(* Logix 5000 project; controller MV vendor 1 type 14 code 217 rev 31.11; software revision 31.00; part 49 of 53 *)
(* tags used below, declared in another part *)
   CheckTimeMask : INT;
   CWD : CHECKWORD_FLAGS;
   Delphi_Does_Eng_Func : BOOL;
   MV_MV10R : PlantItem;   // MV10R
   MV_MV11R : PlantItem;   // MV11R
   MV_MV12R : PlantItem;   // MV12R
   MV_MV13R : PlantItem;   // MV13R
   MV_MV14R : PlantItem;   // MV14R
   MV_MV15R : PlantItem;   // MV15R
   MV_MV16R : PlantItem;   // MV16R
   MV_MV17R : PlantItem;   // MV17R
   MV_MV18R : PlantItem;   // MV18R
   MV_MV19R : PlantItem;   // MV19R
   MV_MV1R : PlantItem;   // MV1R
   MV_MV20R : PlantItem;   // MV20R
   MV_MV21R : PlantItem;   // MV21R
   MV_MV22R : PlantItem;   // MV22R
   MV_MV23R : PlantItem;   // MV23R
   MV_MV2R : PlantItem;   // MV2R
   MV_MV30R : PlantItem;   // MV30R
   MV_MV31R : PlantItem;   // MV31R
   MV_MV32R : PlantItem;   // MV32R
   MV_MV33R : PlantItem;   // MV33R
   MV_MV34R : PlantItem;   // MV34R
   MV_MV35R : PlantItem;   // MV35R
   MV_MV3R : PlantItem;   // MV3R
   MV_MV4R : PlantItem;   // MV4R
   MV_MV5R : PlantItem;   // MV5R
   MV_MV6R : PlantItem;   // MV6R
   MV_MV8R : PlantItem;   // MV8R
   MV_MV9R : PlantItem;   // MV9R
   MV_N255 : DINT[255];   // Old Format Checkwords To Keep Delphi Indicating Status Correctly.
   TempChecktime : DINT;
(* MV_Common, continued *)

   48: [XIC(Delphi_Does_Eng_Func) [[XIC(MV_N255[39].8) [OTL(MV_MV8R.CW.[CWD.MANUAL]) ,XIC(MV_N255[39].9) OTL(MV_MV8R.CW.[CWD.MANDRV]) ,XIO(MV_N255[39].9) OTU(MV_MV8R.CW.[CWD.MANDRV]) ] ,XIO(MV_N255[39].8) [OTU(MV_MV8R.CW.[CWD.MANUAL]) ,[XIC(MV_MV8R.CW.[CWD.OUTPUT]) OTL(MV_N255[39].9) ,XIO(MV_MV8R.CW.[CWD.OUTPUT]) OTU(MV_N255[39].9) ] ] ] ,[XIC(MV_N255[39].13) OTL(MV_MV8R.CW.[CWD.CHECKOFF]) ,XIO(MV_N255[39].13) OTU(MV_MV8R.CW.[CWD.CHECKOFF]) ] ] ,XIO(Delphi_Does_Eng_Func) [[XIC(MV_MV8R.CW.[CWD.MANUAL]) OTL(MV_N255[39].8) ,XIO(MV_MV8R.CW.[CWD.MANUAL]) OTU(MV_N255[39].8) ] ,[XIC(MV_MV8R.CW.[CWD.CHECKOFF]) OTL(MV_N255[39].13) ,XIO(MV_MV8R.CW.[CWD.CHECKOFF]) OTU(MV_N255[39].13) ] ,[XIC(MV_MV8R.CW.[CWD.OUTPUT]) OTL(MV_N255[39].9) ,XIO(MV_MV8R.CW.[CWD.OUTPUT]) OTU(MV_N255[39].9) ] ] ,XIC(MV_MV8R.CW.[CWD.RUNFB]) OTE(MV_N255[39].10) ,XIO(MV_MV8R.CW.[CWD.RUNFB]) OTE(MV_N255[39].11) ,XIC(MV_MV8R.CW.[CWD.FAULT]) OTE(MV_N255[39].15) ];
   49: [XIC(Delphi_Does_Eng_Func) [[XIC(MV_N255[40].8) [OTL(MV_MV9R.CW.[CWD.MANUAL]) ,XIC(MV_N255[40].9) OTL(MV_MV9R.CW.[CWD.MANDRV]) ,XIO(MV_N255[40].9) OTU(MV_MV9R.CW.[CWD.MANDRV]) ] ,XIO(MV_N255[40].8) [OTU(MV_MV9R.CW.[CWD.MANUAL]) ,[XIC(MV_MV9R.CW.[CWD.OUTPUT]) OTL(MV_N255[40].9) ,XIO(MV_MV9R.CW.[CWD.OUTPUT]) OTU(MV_N255[40].9) ] ] ] ,[XIC(MV_N255[40].13) OTL(MV_MV9R.CW.[CWD.CHECKOFF]) ,XIO(MV_N255[40].13) OTU(MV_MV9R.CW.[CWD.CHECKOFF]) ] ] ,XIO(Delphi_Does_Eng_Func) [[XIC(MV_MV9R.CW.[CWD.MANUAL]) OTL(MV_N255[40].8) ,XIO(MV_MV9R.CW.[CWD.MANUAL]) OTU(MV_N255[40].8) ] ,[XIC(MV_MV9R.CW.[CWD.CHECKOFF]) OTL(MV_N255[40].13) ,XIO(MV_MV9R.CW.[CWD.CHECKOFF]) OTU(MV_N255[40].13) ] ,[XIC(MV_MV9R.CW.[CWD.OUTPUT]) OTL(MV_N255[40].9) ,XIO(MV_MV9R.CW.[CWD.OUTPUT]) OTU(MV_N255[40].9) ] ] ,XIC(MV_MV9R.CW.[CWD.RUNFB]) OTE(MV_N255[40].10) ,XIO(MV_MV9R.CW.[CWD.RUNFB]) OTE(MV_N255[40].11) ,XIC(MV_MV9R.CW.[CWD.FAULT]) OTE(MV_N255[40].15) ];
   50: [XIC(Delphi_Does_Eng_Func) [[XIC(MV_N255[41].8) [OTL(MV_MV10R.CW.[CWD.MANUAL]) ,XIC(MV_N255[41].9) OTL(MV_MV10R.CW.[CWD.MANDRV]) ,XIO(MV_N255[41].9) OTU(MV_MV10R.CW.[CWD.MANDRV]) ] ,XIO(MV_N255[41].8) [OTU(MV_MV10R.CW.[CWD.MANUAL]) ,[XIC(MV_MV10R.CW.[CWD.OUTPUT]) OTL(MV_N255[41].9) ,XIO(MV_MV10R.CW.[CWD.OUTPUT]) OTU(MV_N255[41].9) ] ] ] ,[XIC(MV_N255[41].13) OTL(MV_MV10R.CW.[CWD.CHECKOFF]) ,XIO(MV_N255[41].13) OTU(MV_MV10R.CW.[CWD.CHECKOFF]) ] ] ,XIO(Delphi_Does_Eng_Func) [[XIC(MV_MV10R.CW.[CWD.MANUAL]) OTL(MV_N255[41].8) ,XIO(MV_MV10R.CW.[CWD.MANUAL]) OTU(MV_N255[41].8) ] ,[XIC(MV_MV10R.CW.[CWD.CHECKOFF]) OTL(MV_N255[41].13) ,XIO(MV_MV10R.CW.[CWD.CHECKOFF]) OTU(MV_N255[41].13) ] ,[XIC(MV_MV10R.CW.[CWD.OUTPUT]) OTL(MV_N255[41].9) ,XIO(MV_MV10R.CW.[CWD.OUTPUT]) OTU(MV_N255[41].9) ] ] ,XIC(MV_MV10R.CW.[CWD.RUNFB]) OTE(MV_N255[41].10) ,XIO(MV_MV10R.CW.[CWD.RUNFB]) OTE(MV_N255[41].11) ,XIC(MV_MV10R.CW.[CWD.FAULT]) OTE(MV_N255[41].15) ];
   51: [XIC(Delphi_Does_Eng_Func) [[XIC(MV_N255[42].8) [OTL(MV_MV11R.CW.[CWD.MANUAL]) ,XIC(MV_N255[42].9) OTL(MV_MV11R.CW.[CWD.MANDRV]) ,XIO(MV_N255[42].9) OTU(MV_MV11R.CW.[CWD.MANDRV]) ] ,XIO(MV_N255[42].8) [OTU(MV_MV11R.CW.[CWD.MANUAL]) ,[XIC(MV_MV11R.CW.[CWD.OUTPUT]) OTL(MV_N255[42].9) ,XIO(MV_MV11R.CW.[CWD.OUTPUT]) OTU(MV_N255[42].9) ] ] ] ,[XIC(MV_N255[42].13) OTL(MV_MV11R.CW.[CWD.CHECKOFF]) ,XIO(MV_N255[42].13) OTU(MV_MV11R.CW.[CWD.CHECKOFF]) ] ] ,XIO(Delphi_Does_Eng_Func) [[XIC(MV_MV11R.CW.[CWD.MANUAL]) OTL(MV_N255[42].8) ,XIO(MV_MV11R.CW.[CWD.MANUAL]) OTU(MV_N255[42].8) ] ,[XIC(MV_MV11R.CW.[CWD.CHECKOFF]) OTL(MV_N255[42].13) ,XIO(MV_MV11R.CW.[CWD.CHECKOFF]) OTU(MV_N255[42].13) ] ,[XIC(MV_MV11R.CW.[CWD.OUTPUT]) OTL(MV_N255[42].9) ,XIO(MV_MV11R.CW.[CWD.OUTPUT]) OTU(MV_N255[42].9) ] ] ,XIC(MV_MV11R.CW.[CWD.RUNFB]) OTE(MV_N255[42].10) ,XIO(MV_MV11R.CW.[CWD.RUNFB]) OTE(MV_N255[42].11) ,XIC(MV_MV11R.CW.[CWD.FAULT]) OTE(MV_N255[42].15) ];
   52: [XIC(Delphi_Does_Eng_Func) [[XIC(MV_N255[43].8) [OTL(MV_MV12R.CW.[CWD.MANUAL]) ,XIC(MV_N255[43].9) OTL(MV_MV12R.CW.[CWD.MANDRV]) ,XIO(MV_N255[43].9) OTU(MV_MV12R.CW.[CWD.MANDRV]) ] ,XIO(MV_N255[43].8) [OTU(MV_MV12R.CW.[CWD.MANUAL]) ,[XIC(MV_MV12R.CW.[CWD.OUTPUT]) OTL(MV_N255[43].9) ,XIO(MV_MV12R.CW.[CWD.OUTPUT]) OTU(MV_N255[43].9) ] ] ] ,[XIC(MV_N255[43].13) OTL(MV_MV12R.CW.[CWD.CHECKOFF]) ,XIO(MV_N255[43].13) OTU(MV_MV12R.CW.[CWD.CHECKOFF]) ] ] ,XIO(Delphi_Does_Eng_Func) [[XIC(MV_MV12R.CW.[CWD.MANUAL]) OTL(MV_N255[43].8) ,XIO(MV_MV12R.CW.[CWD.MANUAL]) OTU(MV_N255[43].8) ] ,[XIC(MV_MV12R.CW.[CWD.CHECKOFF]) OTL(MV_N255[43].13) ,XIO(MV_MV12R.CW.[CWD.CHECKOFF]) OTU(MV_N255[43].13) ] ,[XIC(MV_MV12R.CW.[CWD.OUTPUT]) OTL(MV_N255[43].9) ,XIO(MV_MV12R.CW.[CWD.OUTPUT]) OTU(MV_N255[43].9) ] ] ,XIC(MV_MV12R.CW.[CWD.RUNFB]) OTE(MV_N255[43].10) ,XIO(MV_MV12R.CW.[CWD.RUNFB]) OTE(MV_N255[43].11) ,XIC(MV_MV12R.CW.[CWD.FAULT]) OTE(MV_N255[43].15) ];
   53: [XIC(Delphi_Does_Eng_Func) [[XIC(MV_N255[44].8) [OTL(MV_MV13R.CW.[CWD.MANUAL]) ,XIC(MV_N255[44].9) OTL(MV_MV13R.CW.[CWD.MANDRV]) ,XIO(MV_N255[44].9) OTU(MV_MV13R.CW.[CWD.MANDRV]) ] ,XIO(MV_N255[44].8) [OTU(MV_MV13R.CW.[CWD.MANUAL]) ,[XIC(MV_MV13R.CW.[CWD.OUTPUT]) OTL(MV_N255[44].9) ,XIO(MV_MV13R.CW.[CWD.OUTPUT]) OTU(MV_N255[44].9) ] ] ] ,[XIC(MV_N255[44].13) OTL(MV_MV13R.CW.[CWD.CHECKOFF]) ,XIO(MV_N255[44].13) OTU(MV_MV13R.CW.[CWD.CHECKOFF]) ] ] ,XIO(Delphi_Does_Eng_Func) [[XIC(MV_MV13R.CW.[CWD.MANUAL]) OTL(MV_N255[44].8) ,XIO(MV_MV13R.CW.[CWD.MANUAL]) OTU(MV_N255[44].8) ] ,[XIC(MV_MV13R.CW.[CWD.CHECKOFF]) OTL(MV_N255[44].13) ,XIO(MV_MV13R.CW.[CWD.CHECKOFF]) OTU(MV_N255[44].13) ] ,[XIC(MV_MV13R.CW.[CWD.OUTPUT]) OTL(MV_N255[44].9) ,XIO(MV_MV13R.CW.[CWD.OUTPUT]) OTU(MV_N255[44].9) ] ] ,XIC(MV_MV13R.CW.[CWD.RUNFB]) OTE(MV_N255[44].10) ,XIO(MV_MV13R.CW.[CWD.RUNFB]) OTE(MV_N255[44].11) ,XIC(MV_MV13R.CW.[CWD.FAULT]) OTE(MV_N255[44].15) ];
   54: [XIC(Delphi_Does_Eng_Func) [[XIC(MV_N255[45].8) [OTL(MV_MV14R.CW.[CWD.MANUAL]) ,XIC(MV_N255[45].9) OTL(MV_MV14R.CW.[CWD.MANDRV]) ,XIO(MV_N255[45].9) OTU(MV_MV14R.CW.[CWD.MANDRV]) ] ,XIO(MV_N255[45].8) [OTU(MV_MV14R.CW.[CWD.MANUAL]) ,[XIC(MV_MV14R.CW.[CWD.OUTPUT]) OTL(MV_N255[45].9) ,XIO(MV_MV14R.CW.[CWD.OUTPUT]) OTU(MV_N255[45].9) ] ] ] ,[XIC(MV_N255[45].13) OTL(MV_MV14R.CW.[CWD.CHECKOFF]) ,XIO(MV_N255[45].13) OTU(MV_MV14R.CW.[CWD.CHECKOFF]) ] ] ,XIO(Delphi_Does_Eng_Func) [[XIC(MV_MV14R.CW.[CWD.MANUAL]) OTL(MV_N255[45].8) ,XIO(MV_MV14R.CW.[CWD.MANUAL]) OTU(MV_N255[45].8) ] ,[XIC(MV_MV14R.CW.[CWD.CHECKOFF]) OTL(MV_N255[45].13) ,XIO(MV_MV14R.CW.[CWD.CHECKOFF]) OTU(MV_N255[45].13) ] ,[XIC(MV_MV14R.CW.[CWD.OUTPUT]) OTL(MV_N255[45].9) ,XIO(MV_MV14R.CW.[CWD.OUTPUT]) OTU(MV_N255[45].9) ] ] ,XIC(MV_MV14R.CW.[CWD.RUNFB]) OTE(MV_N255[45].10) ,XIO(MV_MV14R.CW.[CWD.RUNFB]) OTE(MV_N255[45].11) ,XIC(MV_MV14R.CW.[CWD.FAULT]) OTE(MV_N255[45].15) ];
   55: [XIC(Delphi_Does_Eng_Func) [[XIC(MV_N255[46].8) [OTL(MV_MV15R.CW.[CWD.MANUAL]) ,XIC(MV_N255[46].9) OTL(MV_MV15R.CW.[CWD.MANDRV]) ,XIO(MV_N255[46].9) OTU(MV_MV15R.CW.[CWD.MANDRV]) ] ,XIO(MV_N255[46].8) [OTU(MV_MV15R.CW.[CWD.MANUAL]) ,[XIC(MV_MV15R.CW.[CWD.OUTPUT]) OTL(MV_N255[46].9) ,XIO(MV_MV15R.CW.[CWD.OUTPUT]) OTU(MV_N255[46].9) ] ] ] ,[XIC(MV_N255[46].13) OTL(MV_MV15R.CW.[CWD.CHECKOFF]) ,XIO(MV_N255[46].13) OTU(MV_MV15R.CW.[CWD.CHECKOFF]) ] ] ,XIO(Delphi_Does_Eng_Func) [[XIC(MV_MV15R.CW.[CWD.MANUAL]) OTL(MV_N255[46].8) ,XIO(MV_MV15R.CW.[CWD.MANUAL]) OTU(MV_N255[46].8) ] ,[XIC(MV_MV15R.CW.[CWD.CHECKOFF]) OTL(MV_N255[46].13) ,XIO(MV_MV15R.CW.[CWD.CHECKOFF]) OTU(MV_N255[46].13) ] ,[XIC(MV_MV15R.CW.[CWD.OUTPUT]) OTL(MV_N255[46].9) ,XIO(MV_MV15R.CW.[CWD.OUTPUT]) OTU(MV_N255[46].9) ] ] ,XIC(MV_MV15R.CW.[CWD.RUNFB]) OTE(MV_N255[46].10) ,XIO(MV_MV15R.CW.[CWD.RUNFB]) OTE(MV_N255[46].11) ,XIC(MV_MV15R.CW.[CWD.FAULT]) OTE(MV_N255[46].15) ];
   56: [XIC(Delphi_Does_Eng_Func) [[XIC(MV_N255[47].8) [OTL(MV_MV16R.CW.[CWD.MANUAL]) ,XIC(MV_N255[47].9) OTL(MV_MV16R.CW.[CWD.MANDRV]) ,XIO(MV_N255[47].9) OTU(MV_MV16R.CW.[CWD.MANDRV]) ] ,XIO(MV_N255[47].8) [OTU(MV_MV16R.CW.[CWD.MANUAL]) ,[XIC(MV_MV16R.CW.[CWD.OUTPUT]) OTL(MV_N255[47].9) ,XIO(MV_MV16R.CW.[CWD.OUTPUT]) OTU(MV_N255[47].9) ] ] ] ,[XIC(MV_N255[47].13) OTL(MV_MV16R.CW.[CWD.CHECKOFF]) ,XIO(MV_N255[47].13) OTU(MV_MV16R.CW.[CWD.CHECKOFF]) ] ] ,XIO(Delphi_Does_Eng_Func) [[XIC(MV_MV16R.CW.[CWD.MANUAL]) OTL(MV_N255[47].8) ,XIO(MV_MV16R.CW.[CWD.MANUAL]) OTU(MV_N255[47].8) ] ,[XIC(MV_MV16R.CW.[CWD.CHECKOFF]) OTL(MV_N255[47].13) ,XIO(MV_MV16R.CW.[CWD.CHECKOFF]) OTU(MV_N255[47].13) ] ,[XIC(MV_MV16R.CW.[CWD.OUTPUT]) OTL(MV_N255[47].9) ,XIO(MV_MV16R.CW.[CWD.OUTPUT]) OTU(MV_N255[47].9) ] ] ,XIC(MV_MV16R.CW.[CWD.RUNFB]) OTE(MV_N255[47].10) ,XIO(MV_MV16R.CW.[CWD.RUNFB]) OTE(MV_N255[47].11) ,XIC(MV_MV16R.CW.[CWD.FAULT]) OTE(MV_N255[47].15) ];
   57: [XIC(Delphi_Does_Eng_Func) [[XIC(MV_N255[48].8) [OTL(MV_MV17R.CW.[CWD.MANUAL]) ,XIC(MV_N255[48].9) OTL(MV_MV17R.CW.[CWD.MANDRV]) ,XIO(MV_N255[48].9) OTU(MV_MV17R.CW.[CWD.MANDRV]) ] ,XIO(MV_N255[48].8) [OTU(MV_MV17R.CW.[CWD.MANUAL]) ,[XIC(MV_MV17R.CW.[CWD.OUTPUT]) OTL(MV_N255[48].9) ,XIO(MV_MV17R.CW.[CWD.OUTPUT]) OTU(MV_N255[48].9) ] ] ] ,[XIC(MV_N255[48].13) OTL(MV_MV17R.CW.[CWD.CHECKOFF]) ,XIO(MV_N255[48].13) OTU(MV_MV17R.CW.[CWD.CHECKOFF]) ] ] ,XIO(Delphi_Does_Eng_Func) [[XIC(MV_MV17R.CW.[CWD.MANUAL]) OTL(MV_N255[48].8) ,XIO(MV_MV17R.CW.[CWD.MANUAL]) OTU(MV_N255[48].8) ] ,[XIC(MV_MV17R.CW.[CWD.CHECKOFF]) OTL(MV_N255[48].13) ,XIO(MV_MV17R.CW.[CWD.CHECKOFF]) OTU(MV_N255[48].13) ] ,[XIC(MV_MV17R.CW.[CWD.OUTPUT]) OTL(MV_N255[48].9) ,XIO(MV_MV17R.CW.[CWD.OUTPUT]) OTU(MV_N255[48].9) ] ] ,XIC(MV_MV17R.CW.[CWD.RUNFB]) OTE(MV_N255[48].10) ,XIO(MV_MV17R.CW.[CWD.RUNFB]) OTE(MV_N255[48].11) ,XIC(MV_MV17R.CW.[CWD.FAULT]) OTE(MV_N255[48].15) ];
   58: [XIC(Delphi_Does_Eng_Func) [[XIC(MV_N255[49].8) [OTL(MV_MV18R.CW.[CWD.MANUAL]) ,XIC(MV_N255[49].9) OTL(MV_MV18R.CW.[CWD.MANDRV]) ,XIO(MV_N255[49].9) OTU(MV_MV18R.CW.[CWD.MANDRV]) ] ,XIO(MV_N255[49].8) [OTU(MV_MV18R.CW.[CWD.MANUAL]) ,[XIC(MV_MV18R.CW.[CWD.OUTPUT]) OTL(MV_N255[49].9) ,XIO(MV_MV18R.CW.[CWD.OUTPUT]) OTU(MV_N255[49].9) ] ] ] ,[XIC(MV_N255[49].13) OTL(MV_MV18R.CW.[CWD.CHECKOFF]) ,XIO(MV_N255[49].13) OTU(MV_MV18R.CW.[CWD.CHECKOFF]) ] ] ,XIO(Delphi_Does_Eng_Func) [[XIC(MV_MV18R.CW.[CWD.MANUAL]) OTL(MV_N255[49].8) ,XIO(MV_MV18R.CW.[CWD.MANUAL]) OTU(MV_N255[49].8) ] ,[XIC(MV_MV18R.CW.[CWD.CHECKOFF]) OTL(MV_N255[49].13) ,XIO(MV_MV18R.CW.[CWD.CHECKOFF]) OTU(MV_N255[49].13) ] ,[XIC(MV_MV18R.CW.[CWD.OUTPUT]) OTL(MV_N255[49].9) ,XIO(MV_MV18R.CW.[CWD.OUTPUT]) OTU(MV_N255[49].9) ] ] ,XIC(MV_MV18R.CW.[CWD.RUNFB]) OTE(MV_N255[49].10) ,XIO(MV_MV18R.CW.[CWD.RUNFB]) OTE(MV_N255[49].11) ,XIC(MV_MV18R.CW.[CWD.FAULT]) OTE(MV_N255[49].15) ];
   59: [XIC(Delphi_Does_Eng_Func) [[XIC(MV_N255[50].8) [OTL(MV_MV19R.CW.[CWD.MANUAL]) ,XIC(MV_N255[50].9) OTL(MV_MV19R.CW.[CWD.MANDRV]) ,XIO(MV_N255[50].9) OTU(MV_MV19R.CW.[CWD.MANDRV]) ] ,XIO(MV_N255[50].8) [OTU(MV_MV19R.CW.[CWD.MANUAL]) ,[XIC(MV_MV19R.CW.[CWD.OUTPUT]) OTL(MV_N255[50].9) ,XIO(MV_MV19R.CW.[CWD.OUTPUT]) OTU(MV_N255[50].9) ] ] ] ,[XIC(MV_N255[50].13) OTL(MV_MV19R.CW.[CWD.CHECKOFF]) ,XIO(MV_N255[50].13) OTU(MV_MV19R.CW.[CWD.CHECKOFF]) ] ] ,XIO(Delphi_Does_Eng_Func) [[XIC(MV_MV19R.CW.[CWD.MANUAL]) OTL(MV_N255[50].8) ,XIO(MV_MV19R.CW.[CWD.MANUAL]) OTU(MV_N255[50].8) ] ,[XIC(MV_MV19R.CW.[CWD.CHECKOFF]) OTL(MV_N255[50].13) ,XIO(MV_MV19R.CW.[CWD.CHECKOFF]) OTU(MV_N255[50].13) ] ,[XIC(MV_MV19R.CW.[CWD.OUTPUT]) OTL(MV_N255[50].9) ,XIO(MV_MV19R.CW.[CWD.OUTPUT]) OTU(MV_N255[50].9) ] ] ,XIC(MV_MV19R.CW.[CWD.RUNFB]) OTE(MV_N255[50].10) ,XIO(MV_MV19R.CW.[CWD.RUNFB]) OTE(MV_N255[50].11) ,XIC(MV_MV19R.CW.[CWD.FAULT]) OTE(MV_N255[50].15) ];
   60: [XIC(Delphi_Does_Eng_Func) [[XIC(MV_N255[51].8) [OTL(MV_MV30R.CW.[CWD.MANUAL]) ,XIC(MV_N255[51].9) OTL(MV_MV30R.CW.[CWD.MANDRV]) ,XIO(MV_N255[51].9) OTU(MV_MV30R.CW.[CWD.MANDRV]) ] ,XIO(MV_N255[51].8) [OTU(MV_MV30R.CW.[CWD.MANUAL]) ,[XIC(MV_MV30R.CW.[CWD.OUTPUT]) OTL(MV_N255[51].9) ,XIO(MV_MV30R.CW.[CWD.OUTPUT]) OTU(MV_N255[51].9) ] ] ] ,[XIC(MV_N255[51].13) OTL(MV_MV30R.CW.[CWD.CHECKOFF]) ,XIO(MV_N255[51].13) OTU(MV_MV30R.CW.[CWD.CHECKOFF]) ] ] ,XIO(Delphi_Does_Eng_Func) [[XIC(MV_MV30R.CW.[CWD.MANUAL]) OTL(MV_N255[51].8) ,XIO(MV_MV30R.CW.[CWD.MANUAL]) OTU(MV_N255[51].8) ] ,[XIC(MV_MV30R.CW.[CWD.CHECKOFF]) OTL(MV_N255[51].13) ,XIO(MV_MV30R.CW.[CWD.CHECKOFF]) OTU(MV_N255[51].13) ] ,[XIC(MV_MV30R.CW.[CWD.OUTPUT]) OTL(MV_N255[51].9) ,XIO(MV_MV30R.CW.[CWD.OUTPUT]) OTU(MV_N255[51].9) ] ] ,XIC(MV_MV30R.CW.[CWD.RUNFB]) OTE(MV_N255[51].10) ,XIO(MV_MV30R.CW.[CWD.RUNFB]) OTE(MV_N255[51].11) ,XIC(MV_MV30R.CW.[CWD.FAULT]) OTE(MV_N255[51].15) ];
   61: [XIC(Delphi_Does_Eng_Func) [[XIC(MV_N255[52].8) [OTL(MV_MV31R.CW.[CWD.MANUAL]) ,XIC(MV_N255[52].9) OTL(MV_MV31R.CW.[CWD.MANDRV]) ,XIO(MV_N255[52].9) OTU(MV_MV31R.CW.[CWD.MANDRV]) ] ,XIO(MV_N255[52].8) [OTU(MV_MV31R.CW.[CWD.MANUAL]) ,[XIC(MV_MV31R.CW.[CWD.OUTPUT]) OTL(MV_N255[52].9) ,XIO(MV_MV31R.CW.[CWD.OUTPUT]) OTU(MV_N255[52].9) ] ] ] ,[XIC(MV_N255[52].13) OTL(MV_MV31R.CW.[CWD.CHECKOFF]) ,XIO(MV_N255[52].13) OTU(MV_MV31R.CW.[CWD.CHECKOFF]) ] ] ,XIO(Delphi_Does_Eng_Func) [[XIC(MV_MV31R.CW.[CWD.MANUAL]) OTL(MV_N255[52].8) ,XIO(MV_MV31R.CW.[CWD.MANUAL]) OTU(MV_N255[52].8) ] ,[XIC(MV_MV31R.CW.[CWD.CHECKOFF]) OTL(MV_N255[52].13) ,XIO(MV_MV31R.CW.[CWD.CHECKOFF]) OTU(MV_N255[52].13) ] ,[XIC(MV_MV31R.CW.[CWD.OUTPUT]) OTL(MV_N255[52].9) ,XIO(MV_MV31R.CW.[CWD.OUTPUT]) OTU(MV_N255[52].9) ] ] ,XIC(MV_MV31R.CW.[CWD.RUNFB]) OTE(MV_N255[52].10) ,XIO(MV_MV31R.CW.[CWD.RUNFB]) OTE(MV_N255[52].11) ,XIC(MV_MV31R.CW.[CWD.FAULT]) OTE(MV_N255[52].15) ];
   62: [XIC(Delphi_Does_Eng_Func) [[XIC(MV_N255[53].8) [OTL(MV_MV32R.CW.[CWD.MANUAL]) ,XIC(MV_N255[53].9) OTL(MV_MV32R.CW.[CWD.MANDRV]) ,XIO(MV_N255[53].9) OTU(MV_MV32R.CW.[CWD.MANDRV]) ] ,XIO(MV_N255[53].8) [OTU(MV_MV32R.CW.[CWD.MANUAL]) ,[XIC(MV_MV32R.CW.[CWD.OUTPUT]) OTL(MV_N255[53].9) ,XIO(MV_MV32R.CW.[CWD.OUTPUT]) OTU(MV_N255[53].9) ] ] ] ,[XIC(MV_N255[53].13) OTL(MV_MV32R.CW.[CWD.CHECKOFF]) ,XIO(MV_N255[53].13) OTU(MV_MV32R.CW.[CWD.CHECKOFF]) ] ] ,XIO(Delphi_Does_Eng_Func) [[XIC(MV_MV32R.CW.[CWD.MANUAL]) OTL(MV_N255[53].8) ,XIO(MV_MV32R.CW.[CWD.MANUAL]) OTU(MV_N255[53].8) ] ,[XIC(MV_MV32R.CW.[CWD.CHECKOFF]) OTL(MV_N255[53].13) ,XIO(MV_MV32R.CW.[CWD.CHECKOFF]) OTU(MV_N255[53].13) ] ,[XIC(MV_MV32R.CW.[CWD.OUTPUT]) OTL(MV_N255[53].9) ,XIO(MV_MV32R.CW.[CWD.OUTPUT]) OTU(MV_N255[53].9) ] ] ,XIC(MV_MV32R.CW.[CWD.RUNFB]) OTE(MV_N255[53].10) ,XIO(MV_MV32R.CW.[CWD.RUNFB]) OTE(MV_N255[53].11) ,XIC(MV_MV32R.CW.[CWD.FAULT]) OTE(MV_N255[53].15) ];
   63: [XIC(Delphi_Does_Eng_Func) [[XIC(MV_N255[54].8) [OTL(MV_MV33R.CW.[CWD.MANUAL]) ,XIC(MV_N255[54].9) OTL(MV_MV33R.CW.[CWD.MANDRV]) ,XIO(MV_N255[54].9) OTU(MV_MV33R.CW.[CWD.MANDRV]) ] ,XIO(MV_N255[54].8) [OTU(MV_MV33R.CW.[CWD.MANUAL]) ,[XIC(MV_MV33R.CW.[CWD.OUTPUT]) OTL(MV_N255[54].9) ,XIO(MV_MV33R.CW.[CWD.OUTPUT]) OTU(MV_N255[54].9) ] ] ] ,[XIC(MV_N255[54].13) OTL(MV_MV33R.CW.[CWD.CHECKOFF]) ,XIO(MV_N255[54].13) OTU(MV_MV33R.CW.[CWD.CHECKOFF]) ] ] ,XIO(Delphi_Does_Eng_Func) [[XIC(MV_MV33R.CW.[CWD.MANUAL]) OTL(MV_N255[54].8) ,XIO(MV_MV33R.CW.[CWD.MANUAL]) OTU(MV_N255[54].8) ] ,[XIC(MV_MV33R.CW.[CWD.CHECKOFF]) OTL(MV_N255[54].13) ,XIO(MV_MV33R.CW.[CWD.CHECKOFF]) OTU(MV_N255[54].13) ] ,[XIC(MV_MV33R.CW.[CWD.OUTPUT]) OTL(MV_N255[54].9) ,XIO(MV_MV33R.CW.[CWD.OUTPUT]) OTU(MV_N255[54].9) ] ] ,XIC(MV_MV33R.CW.[CWD.RUNFB]) OTE(MV_N255[54].10) ,XIO(MV_MV33R.CW.[CWD.RUNFB]) OTE(MV_N255[54].11) ,XIC(MV_MV33R.CW.[CWD.FAULT]) OTE(MV_N255[54].15) ];
   64: [XIC(Delphi_Does_Eng_Func) [[XIC(MV_N255[55].8) [OTL(MV_MV34R.CW.[CWD.MANUAL]) ,XIC(MV_N255[55].9) OTL(MV_MV34R.CW.[CWD.MANDRV]) ,XIO(MV_N255[55].9) OTU(MV_MV34R.CW.[CWD.MANDRV]) ] ,XIO(MV_N255[55].8) [OTU(MV_MV34R.CW.[CWD.MANUAL]) ,[XIC(MV_MV34R.CW.[CWD.OUTPUT]) OTL(MV_N255[55].9) ,XIO(MV_MV34R.CW.[CWD.OUTPUT]) OTU(MV_N255[55].9) ] ] ] ,[XIC(MV_N255[55].13) OTL(MV_MV34R.CW.[CWD.CHECKOFF]) ,XIO(MV_N255[55].13) OTU(MV_MV34R.CW.[CWD.CHECKOFF]) ] ] ,XIO(Delphi_Does_Eng_Func) [[XIC(MV_MV34R.CW.[CWD.MANUAL]) OTL(MV_N255[55].8) ,XIO(MV_MV34R.CW.[CWD.MANUAL]) OTU(MV_N255[55].8) ] ,[XIC(MV_MV34R.CW.[CWD.CHECKOFF]) OTL(MV_N255[55].13) ,XIO(MV_MV34R.CW.[CWD.CHECKOFF]) OTU(MV_N255[55].13) ] ,[XIC(MV_MV34R.CW.[CWD.OUTPUT]) OTL(MV_N255[55].9) ,XIO(MV_MV34R.CW.[CWD.OUTPUT]) OTU(MV_N255[55].9) ] ] ,XIC(MV_MV34R.CW.[CWD.RUNFB]) OTE(MV_N255[55].10) ,XIO(MV_MV34R.CW.[CWD.RUNFB]) OTE(MV_N255[55].11) ,XIC(MV_MV34R.CW.[CWD.FAULT]) OTE(MV_N255[55].15) ];
   65: [XIC(Delphi_Does_Eng_Func) [[XIC(MV_N255[56].8) [OTL(MV_MV35R.CW.[CWD.MANUAL]) ,XIC(MV_N255[56].9) OTL(MV_MV35R.CW.[CWD.MANDRV]) ,XIO(MV_N255[56].9) OTU(MV_MV35R.CW.[CWD.MANDRV]) ] ,XIO(MV_N255[56].8) [OTU(MV_MV35R.CW.[CWD.MANUAL]) ,[XIC(MV_MV35R.CW.[CWD.OUTPUT]) OTL(MV_N255[56].9) ,XIO(MV_MV35R.CW.[CWD.OUTPUT]) OTU(MV_N255[56].9) ] ] ] ,[XIC(MV_N255[56].13) OTL(MV_MV35R.CW.[CWD.CHECKOFF]) ,XIO(MV_N255[56].13) OTU(MV_MV35R.CW.[CWD.CHECKOFF]) ] ] ,XIO(Delphi_Does_Eng_Func) [[XIC(MV_MV35R.CW.[CWD.MANUAL]) OTL(MV_N255[56].8) ,XIO(MV_MV35R.CW.[CWD.MANUAL]) OTU(MV_N255[56].8) ] ,[XIC(MV_MV35R.CW.[CWD.CHECKOFF]) OTL(MV_N255[56].13) ,XIO(MV_MV35R.CW.[CWD.CHECKOFF]) OTU(MV_N255[56].13) ] ,[XIC(MV_MV35R.CW.[CWD.OUTPUT]) OTL(MV_N255[56].9) ,XIO(MV_MV35R.CW.[CWD.OUTPUT]) OTU(MV_N255[56].9) ] ] ,XIC(MV_MV35R.CW.[CWD.RUNFB]) OTE(MV_N255[56].10) ,XIO(MV_MV35R.CW.[CWD.RUNFB]) OTE(MV_N255[56].11) ,XIC(MV_MV35R.CW.[CWD.FAULT]) OTE(MV_N255[56].15) ];
   66: [XIC(Delphi_Does_Eng_Func) [[XIC(MV_N255[57].8) [OTL(MV_MV20R.CW.[CWD.MANUAL]) ,XIC(MV_N255[57].9) OTL(MV_MV20R.CW.[CWD.MANDRV]) ,XIO(MV_N255[57].9) OTU(MV_MV20R.CW.[CWD.MANDRV]) ] ,XIO(MV_N255[57].8) [OTU(MV_MV20R.CW.[CWD.MANUAL]) ,[XIC(MV_MV20R.CW.[CWD.OUTPUT]) OTL(MV_N255[57].9) ,XIO(MV_MV20R.CW.[CWD.OUTPUT]) OTU(MV_N255[57].9) ] ] ] ,[XIC(MV_N255[57].13) OTL(MV_MV20R.CW.[CWD.CHECKOFF]) ,XIO(MV_N255[57].13) OTU(MV_MV20R.CW.[CWD.CHECKOFF]) ] ] ,XIO(Delphi_Does_Eng_Func) [[XIC(MV_MV20R.CW.[CWD.MANUAL]) OTL(MV_N255[57].8) ,XIO(MV_MV20R.CW.[CWD.MANUAL]) OTU(MV_N255[57].8) ] ,[XIC(MV_MV20R.CW.[CWD.CHECKOFF]) OTL(MV_N255[57].13) ,XIO(MV_MV20R.CW.[CWD.CHECKOFF]) OTU(MV_N255[57].13) ] ,[XIC(MV_MV20R.CW.[CWD.OUTPUT]) OTL(MV_N255[57].9) ,XIO(MV_MV20R.CW.[CWD.OUTPUT]) OTU(MV_N255[57].9) ] ] ,XIC(MV_MV20R.CW.[CWD.RUNFB]) OTE(MV_N255[57].10) ,XIO(MV_MV20R.CW.[CWD.RUNFB]) OTE(MV_N255[57].11) ,XIC(MV_MV20R.CW.[CWD.FAULT]) OTE(MV_N255[57].15) ];
   67: [XIC(Delphi_Does_Eng_Func) [[XIC(MV_N255[58].8) [OTL(MV_MV21R.CW.[CWD.MANUAL]) ,XIC(MV_N255[58].9) OTL(MV_MV21R.CW.[CWD.MANDRV]) ,XIO(MV_N255[58].9) OTU(MV_MV21R.CW.[CWD.MANDRV]) ] ,XIO(MV_N255[58].8) [OTU(MV_MV21R.CW.[CWD.MANUAL]) ,[XIC(MV_MV21R.CW.[CWD.OUTPUT]) OTL(MV_N255[58].9) ,XIO(MV_MV21R.CW.[CWD.OUTPUT]) OTU(MV_N255[58].9) ] ] ] ,[XIC(MV_N255[58].13) OTL(MV_MV21R.CW.[CWD.CHECKOFF]) ,XIO(MV_N255[58].13) OTU(MV_MV21R.CW.[CWD.CHECKOFF]) ] ] ,XIO(Delphi_Does_Eng_Func) [[XIC(MV_MV21R.CW.[CWD.MANUAL]) OTL(MV_N255[58].8) ,XIO(MV_MV21R.CW.[CWD.MANUAL]) OTU(MV_N255[58].8) ] ,[XIC(MV_MV21R.CW.[CWD.CHECKOFF]) OTL(MV_N255[58].13) ,XIO(MV_MV21R.CW.[CWD.CHECKOFF]) OTU(MV_N255[58].13) ] ,[XIC(MV_MV21R.CW.[CWD.OUTPUT]) OTL(MV_N255[58].9) ,XIO(MV_MV21R.CW.[CWD.OUTPUT]) OTU(MV_N255[58].9) ] ] ,XIC(MV_MV21R.CW.[CWD.RUNFB]) OTE(MV_N255[58].10) ,XIO(MV_MV21R.CW.[CWD.RUNFB]) OTE(MV_N255[58].11) ,XIC(MV_MV21R.CW.[CWD.FAULT]) OTE(MV_N255[58].15) ];
   68: [XIC(Delphi_Does_Eng_Func) [[XIC(MV_N255[59].8) [OTL(MV_MV22R.CW.[CWD.MANUAL]) ,XIC(MV_N255[59].9) OTL(MV_MV22R.CW.[CWD.MANDRV]) ,XIO(MV_N255[59].9) OTU(MV_MV22R.CW.[CWD.MANDRV]) ] ,XIO(MV_N255[59].8) [OTU(MV_MV22R.CW.[CWD.MANUAL]) ,[XIC(MV_MV22R.CW.[CWD.OUTPUT]) OTL(MV_N255[59].9) ,XIO(MV_MV22R.CW.[CWD.OUTPUT]) OTU(MV_N255[59].9) ] ] ] ,[XIC(MV_N255[59].13) OTL(MV_MV22R.CW.[CWD.CHECKOFF]) ,XIO(MV_N255[59].13) OTU(MV_MV22R.CW.[CWD.CHECKOFF]) ] ] ,XIO(Delphi_Does_Eng_Func) [[XIC(MV_MV22R.CW.[CWD.MANUAL]) OTL(MV_N255[59].8) ,XIO(MV_MV22R.CW.[CWD.MANUAL]) OTU(MV_N255[59].8) ] ,[XIC(MV_MV22R.CW.[CWD.CHECKOFF]) OTL(MV_N255[59].13) ,XIO(MV_MV22R.CW.[CWD.CHECKOFF]) OTU(MV_N255[59].13) ] ,[XIC(MV_MV22R.CW.[CWD.OUTPUT]) OTL(MV_N255[59].9) ,XIO(MV_MV22R.CW.[CWD.OUTPUT]) OTU(MV_N255[59].9) ] ] ,XIC(MV_MV22R.CW.[CWD.RUNFB]) OTE(MV_N255[59].10) ,XIO(MV_MV22R.CW.[CWD.RUNFB]) OTE(MV_N255[59].11) ,XIC(MV_MV22R.CW.[CWD.FAULT]) OTE(MV_N255[59].15) ];
   69: [XIC(Delphi_Does_Eng_Func) [[XIC(MV_N255[60].8) [OTL(MV_MV23R.CW.[CWD.MANUAL]) ,XIC(MV_N255[60].9) OTL(MV_MV23R.CW.[CWD.MANDRV]) ,XIO(MV_N255[60].9) OTU(MV_MV23R.CW.[CWD.MANDRV]) ] ,XIO(MV_N255[60].8) [OTU(MV_MV23R.CW.[CWD.MANUAL]) ,[XIC(MV_MV23R.CW.[CWD.OUTPUT]) OTL(MV_N255[60].9) ,XIO(MV_MV23R.CW.[CWD.OUTPUT]) OTU(MV_N255[60].9) ] ] ] ,[XIC(MV_N255[60].13) OTL(MV_MV23R.CW.[CWD.CHECKOFF]) ,XIO(MV_N255[60].13) OTU(MV_MV23R.CW.[CWD.CHECKOFF]) ] ] ,XIO(Delphi_Does_Eng_Func) [[XIC(MV_MV23R.CW.[CWD.MANUAL]) OTL(MV_N255[60].8) ,XIO(MV_MV23R.CW.[CWD.MANUAL]) OTU(MV_N255[60].8) ] ,[XIC(MV_MV23R.CW.[CWD.CHECKOFF]) OTL(MV_N255[60].13) ,XIO(MV_MV23R.CW.[CWD.CHECKOFF]) OTU(MV_N255[60].13) ] ,[XIC(MV_MV23R.CW.[CWD.OUTPUT]) OTL(MV_N255[60].9) ,XIO(MV_MV23R.CW.[CWD.OUTPUT]) OTU(MV_N255[60].9) ] ] ,XIC(MV_MV23R.CW.[CWD.RUNFB]) OTE(MV_N255[60].10) ,XIO(MV_MV23R.CW.[CWD.RUNFB]) OTE(MV_N255[60].11) ,XIC(MV_MV23R.CW.[CWD.FAULT]) OTE(MV_N255[60].15) ];
   70: XIC(Delphi_Does_Eng_Func)AND(MV_N255[32],CheckTimeMask,TempChecktime)[GRT(TempChecktime,0) DIV(TempChecktime,8,MV_MV1R.CheckTime) ,EQU(TempChecktime,0) OTL(MV_N255[32].6) ];
   71: XIC(Delphi_Does_Eng_Func)AND(MV_N255[33],CheckTimeMask,TempChecktime)[GRT(TempChecktime,0) DIV(TempChecktime,8,MV_MV2R.CheckTime) ,EQU(TempChecktime,0) OTL(MV_N255[33].6) ];
   72: XIC(Delphi_Does_Eng_Func)AND(MV_N255[34],CheckTimeMask,TempChecktime)[GRT(TempChecktime,0) DIV(TempChecktime,8,MV_MV3R.CheckTime) ,EQU(TempChecktime,0) OTL(MV_N255[34].6) ];
   73: XIC(Delphi_Does_Eng_Func)AND(MV_N255[35],CheckTimeMask,TempChecktime)[GRT(TempChecktime,0) DIV(TempChecktime,8,MV_MV4R.CheckTime) ,EQU(TempChecktime,0) OTL(MV_N255[35].6) ];
   74: XIC(Delphi_Does_Eng_Func)AND(MV_N255[36],CheckTimeMask,TempChecktime)[GRT(TempChecktime,0) DIV(TempChecktime,8,MV_MV5R.CheckTime) ,EQU(TempChecktime,0) OTL(MV_N255[36].6) ];
   75: XIC(Delphi_Does_Eng_Func)AND(MV_N255[37],CheckTimeMask,TempChecktime)[GRT(TempChecktime,0) DIV(TempChecktime,8,MV_MV6R.CheckTime) ,EQU(TempChecktime,0) OTL(MV_N255[37].6) ];
